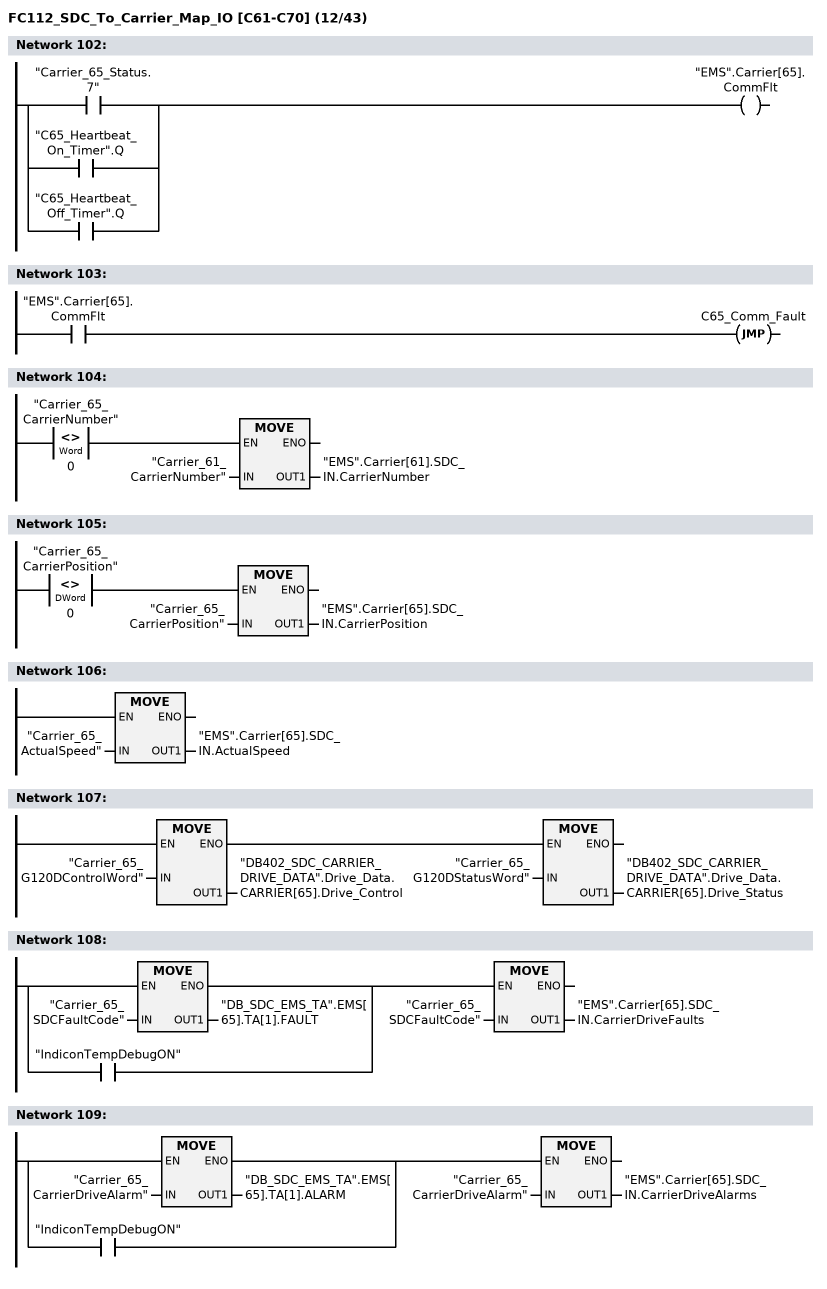
   RUNG wire#powerrail
      Contact( "Carrier_65_Status.7" )
      wire#w1
      Coil( "EMS".Carrier[65].CommFlt )
   END_RUNG
   RUNG wire#powerrail
      Contact( "C65_Heartbeat_On_Timer".Q )
   END_RUNG wire#w1
   RUNG wire#powerrail
      Contact( "C65_Heartbeat_Off_Timer".Q )
   END_RUNG wire#w1
   // the same network as SCL:
   "EMS".Carrier[65].CommFlt := "Carrier_65_Status.7" OR "C65_Heartbeat_On_Timer".Q OR "C65_Heartbeat_Off_Timer".Q;
END_REGION

REGION Network 103
   RUNG wire#powerrail
      Contact( "EMS".Carrier[65].CommFlt )
      JumpCoil( C65_Comm_Fault )
   END_RUNG
   // the same network as SCL:
   IF "EMS".Carrier[65].CommFlt THEN GOTO C65_Comm_Fault; END_IF;
END_REGION

REGION Network 104
   RUNG wire#powerrail
      { S7_Templates := "SrcType := Word" } NE_Contact(in1 := "Carrier_65_CarrierNumber", in2 := 0)
      Move(in := "Carrier_61_CarrierNumber", out1 => "EMS".Carrier[61].SDC_IN.CarrierNumber)
   END_RUNG
   // the same network as SCL:
   IF "Carrier_65_CarrierNumber" <> 0 THEN
       "EMS".Carrier[61].SDC_IN.CarrierNumber := "Carrier_61_CarrierNumber";
   END_IF;
END_REGION

REGION Network 105
   RUNG wire#powerrail
      { S7_Templates := "SrcType := DWord" } NE_Contact(in1 := "Carrier_65_CarrierPosition", in2 := 0)
      Move(in := "Carrier_65_CarrierPosition", out1 => "EMS".Carrier[65].SDC_IN.CarrierPosition)
   END_RUNG
   // the same network as SCL:
   IF "Carrier_65_CarrierPosition" <> 0 THEN
       "EMS".Carrier[65].SDC_IN.CarrierPosition := "Carrier_65_CarrierPosition";
   END_IF;
END_REGION

REGION Network 106
   RUNG wire#powerrail
      Move(in := "Carrier_65_ActualSpeed", out1 => "EMS".Carrier[65].SDC_IN.ActualSpeed)
   END_RUNG
   // the same network as SCL:
   "EMS".Carrier[65].SDC_IN.ActualSpeed := "Carrier_65_ActualSpeed";
END_REGION

REGION Network 107
   RUNG wire#powerrail
      Move(in := "Carrier_65_G120DControlWord", out1 => "DB402_SDC_CARRIER_DRIVE_DATA".Drive_Data.CARRIER[65].Drive_Control)
      Move(in := "Carrier_65_G120DStatusWord", out1 => "DB402_SDC_CARRIER_DRIVE_DATA".Drive_Data.CARRIER[65].Drive_Status)
   END_RUNG
   // the same network as SCL:
   "DB402_SDC_CARRIER_DRIVE_DATA".Drive_Data.CARRIER[65].Drive_Control := "Carrier_65_G120DControlWord";
   "DB402_SDC_CARRIER_DRIVE_DATA".Drive_Data.CARRIER[65].Drive_Status := "Carrier_65_G120DStatusWord";
END_REGION

REGION Network 108
   RUNG wire#powerrail
      Move(in := "Carrier_65_SDCFaultCode", out1 => "DB_SDC_EMS_TA".EMS[65].TA[1].FAULT)
      wire#w1
      Move(in := "Carrier_65_SDCFaultCode", out1 => "EMS".Carrier[65].SDC_IN.CarrierDriveFaults)
   END_RUNG
   RUNG wire#powerrail
      Contact( "IndiconTempDebugON" )
   END_RUNG wire#w1
   // the same network as SCL:
   "DB_SDC_EMS_TA".EMS[65].TA[1].FAULT := "Carrier_65_SDCFaultCode";
   IF TRUE OR "IndiconTempDebugON" THEN
       "EMS".Carrier[65].SDC_IN.CarrierDriveFaults := "Carrier_65_SDCFaultCode";
   END_IF;
END_REGION

REGION Network 109
   RUNG wire#powerrail
      Move(in := "Carrier_65_CarrierDriveAlarm", out1 => "DB_SDC_EMS_TA".EMS[65].TA[1].ALARM)
      wire#w1
      Move(in := "Carrier_65_CarrierDriveAlarm", out1 => "EMS".Carrier[65].SDC_IN.CarrierDriveAlarms)
   END_RUNG
   RUNG wire#powerrail
      Contact( "IndiconTempDebugON" )
   END_RUNG wire#w1
   // the same network as SCL:
   "DB_SDC_EMS_TA".EMS[65].TA[1].ALARM := "Carrier_65_CarrierDriveAlarm";
   IF TRUE OR "IndiconTempDebugON" THEN
       "EMS".Carrier[65].SDC_IN.CarrierDriveAlarms := "Carrier_65_CarrierDriveAlarm";
   END_IF;
END_REGION

REGION Network 110
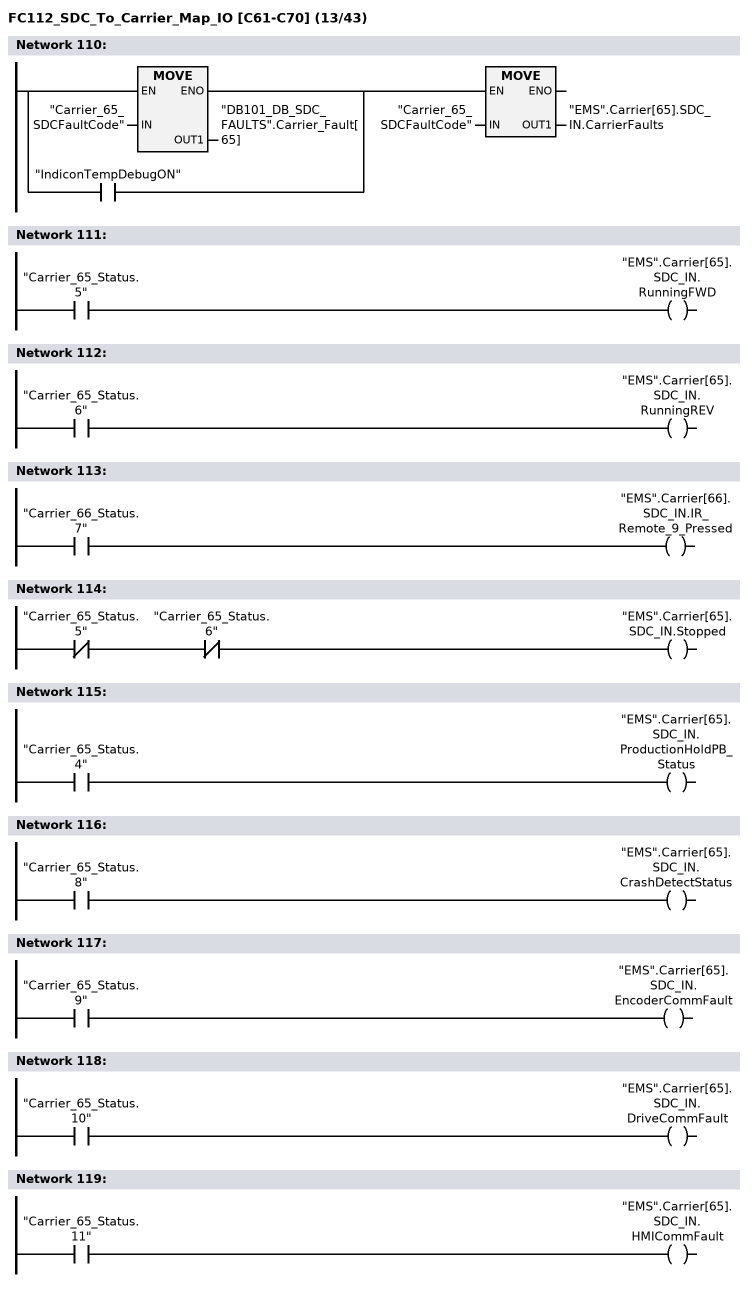
   RUNG wire#powerrail
      Move(in := "Carrier_65_SDCFaultCode", out1 => "DB101_DB_SDC_FAULTS".Carrier_Fault[65])
      wire#w1
      Move(in := "Carrier_65_SDCFaultCode", out1 => "EMS".Carrier[65].SDC_IN.CarrierFaults)
   END_RUNG
   RUNG wire#powerrail
      Contact( "IndiconTempDebugON" )
   END_RUNG wire#w1
   // the same network as SCL:
   "DB101_DB_SDC_FAULTS".Carrier_Fault[65] := "Carrier_65_SDCFaultCode";
   IF TRUE OR "IndiconTempDebugON" THEN
       "EMS".Carrier[65].SDC_IN.CarrierFaults := "Carrier_65_SDCFaultCode";
   END_IF;
END_REGION

REGION Network 111
   RUNG wire#powerrail
      Contact( "Carrier_65_Status.5" )
      Coil( "EMS".Carrier[65].SDC_IN.RunningFWD )
   END_RUNG
   // the same network as SCL:
   "EMS".Carrier[65].SDC_IN.RunningFWD := "Carrier_65_Status.5";
END_REGION

REGION Network 112
   RUNG wire#powerrail
      Contact( "Carrier_65_Status.6" )
      Coil( "EMS".Carrier[65].SDC_IN.RunningREV )
   END_RUNG
   // the same network as SCL:
   "EMS".Carrier[65].SDC_IN.RunningREV := "Carrier_65_Status.6";
END_REGION

REGION Network 113
   RUNG wire#powerrail
      Contact( "Carrier_66_Status.7" )
      Coil( "EMS".Carrier[66].SDC_IN.IR_Remote_9_Pressed )
   END_RUNG
   // the same network as SCL:
   "EMS".Carrier[66].SDC_IN.IR_Remote_9_Pressed := "Carrier_66_Status.7";
END_REGION

REGION Network 114
   RUNG wire#powerrail
      I_Contact( "Carrier_65_Status.5" )
      I_Contact( "Carrier_65_Status.6" )
      Coil( "EMS".Carrier[65].SDC_IN.Stopped )
   END_RUNG
   // the same network as SCL:
   "EMS".Carrier[65].SDC_IN.Stopped := NOT "Carrier_65_Status.5" AND NOT "Carrier_65_Status.6";
END_REGION

REGION Network 115
   RUNG wire#powerrail
      Contact( "Carrier_65_Status.4" )
      Coil( "EMS".Carrier[65].SDC_IN.ProductionHoldPB_Status )
   END_RUNG
   // the same network as SCL:
   "EMS".Carrier[65].SDC_IN.ProductionHoldPB_Status := "Carrier_65_Status.4";
END_REGION

REGION Network 116
   RUNG wire#powerrail
      Contact( "Carrier_65_Status.8" )
      Coil( "EMS".Carrier[65].SDC_IN.CrashDetectStatus )
   END_RUNG
   // the same network as SCL:
   "EMS".Carrier[65].SDC_IN.CrashDetectStatus := "Carrier_65_Status.8";
END_REGION

REGION Network 117
   RUNG wire#powerrail
      Contact( "Carrier_65_Status.9" )
      Coil( "EMS".Carrier[65].SDC_IN.EncoderCommFault )
   END_RUNG
   // the same network as SCL:
   "EMS".Carrier[65].SDC_IN.EncoderCommFault := "Carrier_65_Status.9";
END_REGION

REGION Network 118
   RUNG wire#powerrail
      Contact( "Carrier_65_Status.10" )
      Coil( "EMS".Carrier[65].SDC_IN.DriveCommFault )
   END_RUNG
   // the same network as SCL:
   "EMS".Carrier[65].SDC_IN.DriveCommFault := "Carrier_65_Status.10";
END_REGION

REGION Network 119
   RUNG wire#powerrail
      Contact( "Carrier_65_Status.11" )
      Coil( "EMS".Carrier[65].SDC_IN.HMICommFault )
   END_RUNG
   // the same network as SCL:
   "EMS".Carrier[65].SDC_IN.HMICommFault := "Carrier_65_Status.11";
END_REGION

REGION Network 120
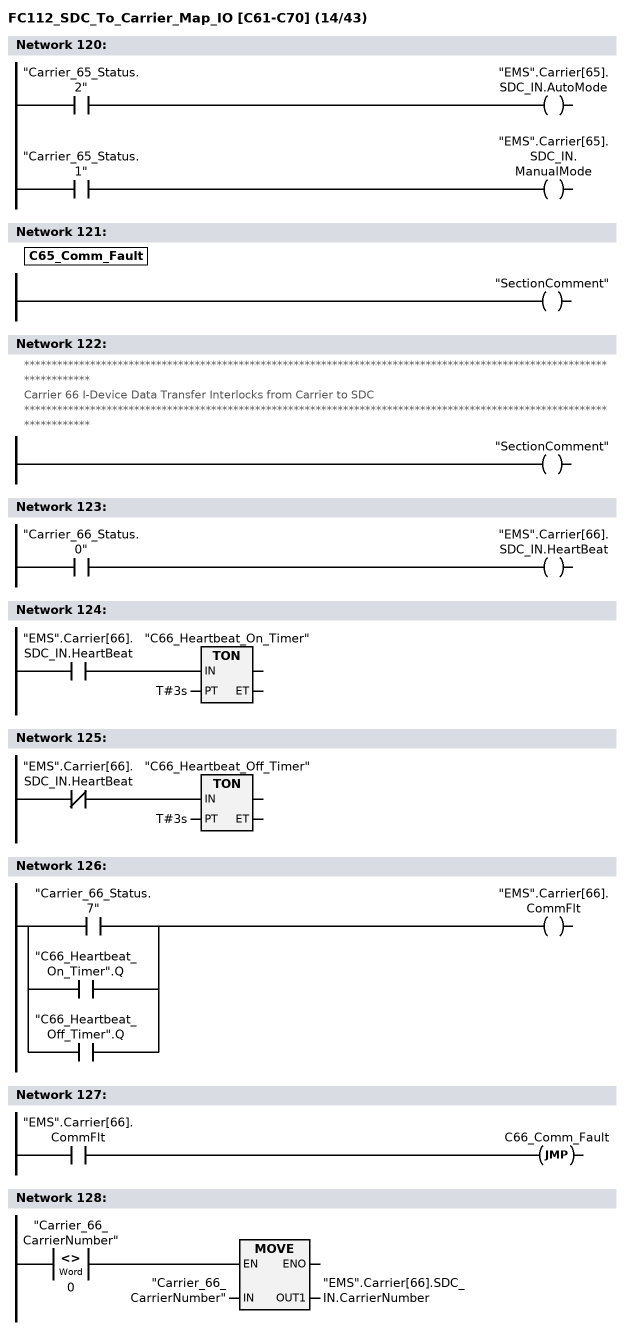
   RUNG wire#powerrail
      Contact( "Carrier_65_Status.2" )
      Coil( "EMS".Carrier[65].SDC_IN.AutoMode )
   END_RUNG
   RUNG wire#powerrail
      Contact( "Carrier_65_Status.1" )
      Coil( "EMS".Carrier[65].SDC_IN.ManualMode )
   END_RUNG
   // the same network as SCL:
   "EMS".Carrier[65].SDC_IN.AutoMode := "Carrier_65_Status.2";
   "EMS".Carrier[65].SDC_IN.ManualMode := "Carrier_65_Status.1";
END_REGION

REGION Network 121
   Label( C65_Comm_Fault )
   RUNG wire#powerrail
      Coil( "SectionComment" )
   END_RUNG
   // the same network as SCL:
   C65_Comm_Fault:
   "SectionComment" := TRUE;
END_REGION

REGION Network 122
   // **********************************************************************************************************************
   // 
   // Carrier 66 I-Device Data Transfer Interlocks from Carrier to SDC
   // 
   // **********************************************************************************************************************
   RUNG wire#powerrail
      Coil( "SectionComment" )
   END_RUNG
   // the same network as SCL:
   "SectionComment" := TRUE;
END_REGION

REGION Network 123
   RUNG wire#powerrail
      Contact( "Carrier_66_Status.0" )
      Coil( "EMS".Carrier[66].SDC_IN.HeartBeat )
   END_RUNG
   // the same network as SCL:
   "EMS".Carrier[66].SDC_IN.HeartBeat := "Carrier_66_Status.0";
END_REGION

REGION Network 124
   "C66_Heartbeat_On_Timer".TON(IN := "EMS".Carrier[66].SDC_IN.HeartBeat, PT := T#3s);
END_REGION

REGION Network 125
   "C66_Heartbeat_Off_Timer".TON(IN := NOT "EMS".Carrier[66].SDC_IN.HeartBeat, PT := T#3s);
END_REGION

REGION Network 126
   RUNG wire#powerrail
      Contact( "Carrier_66_Status.7" )
      wire#w1
      Coil( "EMS".Carrier[66].CommFlt )
   END_RUNG
   RUNG wire#powerrail
      Contact( "C66_Heartbeat_On_Timer".Q )
   END_RUNG wire#w1
   RUNG wire#powerrail
      Contact( "C66_Heartbeat_Off_Timer".Q )
   END_RUNG wire#w1
   // the same network as SCL:
   "EMS".Carrier[66].CommFlt := "Carrier_66_Status.7" OR "C66_Heartbeat_On_Timer".Q OR "C66_Heartbeat_Off_Timer".Q;
END_REGION

REGION Network 127
   RUNG wire#powerrail
      Contact( "EMS".Carrier[66].CommFlt )
      JumpCoil( C66_Comm_Fault )
   END_RUNG
   // the same network as SCL:
   IF "EMS".Carrier[66].CommFlt THEN GOTO C66_Comm_Fault; END_IF;
END_REGION

REGION Network 128
   RUNG wire#powerrail
      { S7_Templates := "SrcType := Word" } NE_Contact(in1 := "Carrier_66_CarrierNumber", in2 := 0)
      Move(in := "Carrier_66_CarrierNumber", out1 => "EMS".Carrier[66].SDC_IN.CarrierNumber)
   END_RUNG
   // the same network as SCL:
   IF "Carrier_66_CarrierNumber" <> 0 THEN
       "EMS".Carrier[66].SDC_IN.CarrierNumber := "Carrier_66_CarrierNumber";
   END_IF;
END_REGION

REGION Network 129
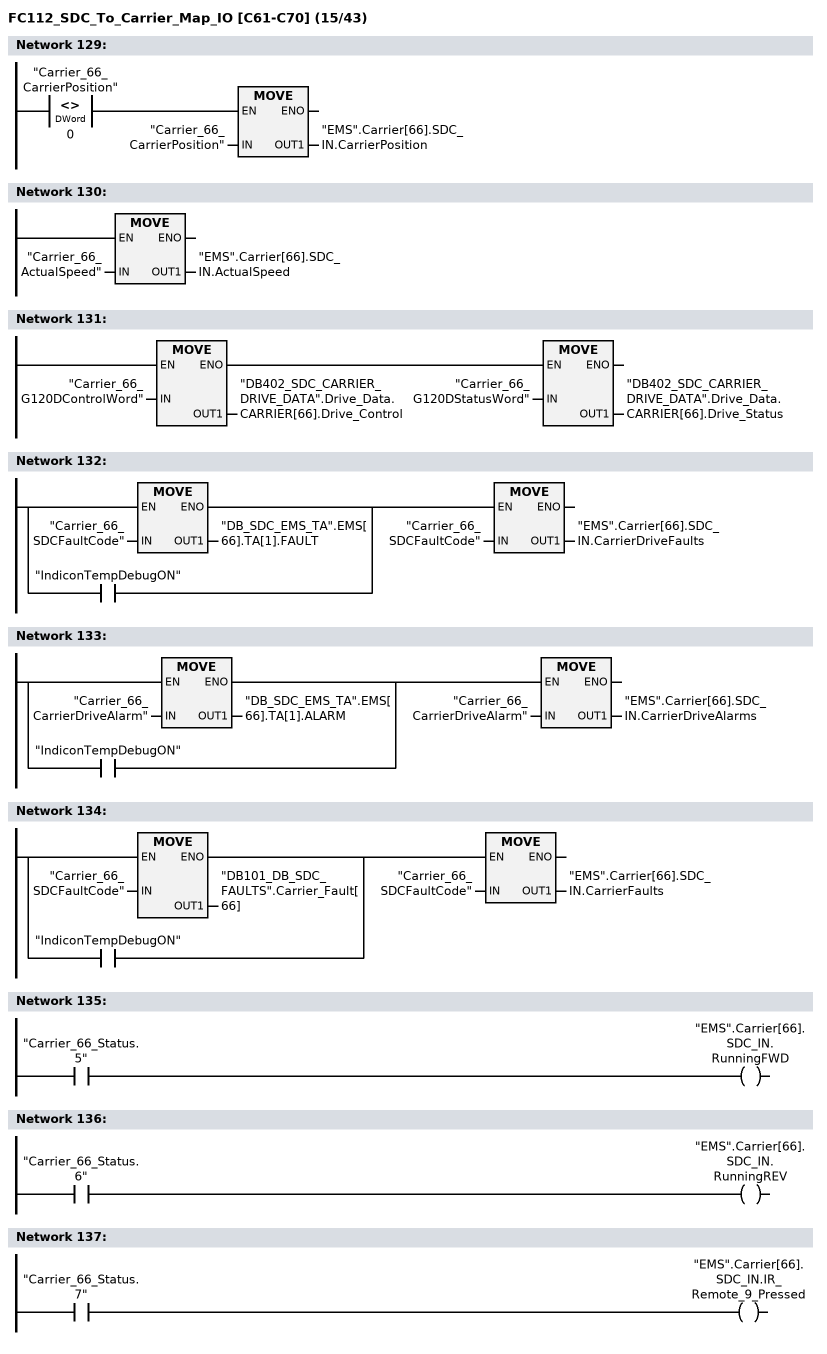
   RUNG wire#powerrail
      { S7_Templates := "SrcType := DWord" } NE_Contact(in1 := "Carrier_66_CarrierPosition", in2 := 0)
      Move(in := "Carrier_66_CarrierPosition", out1 => "EMS".Carrier[66].SDC_IN.CarrierPosition)
   END_RUNG
   // the same network as SCL:
   IF "Carrier_66_CarrierPosition" <> 0 THEN
       "EMS".Carrier[66].SDC_IN.CarrierPosition := "Carrier_66_CarrierPosition";
   END_IF;
END_REGION

REGION Network 130
   RUNG wire#powerrail
      Move(in := "Carrier_66_ActualSpeed", out1 => "EMS".Carrier[66].SDC_IN.ActualSpeed)
   END_RUNG
   // the same network as SCL:
   "EMS".Carrier[66].SDC_IN.ActualSpeed := "Carrier_66_ActualSpeed";
END_REGION

REGION Network 131
   RUNG wire#powerrail
      Move(in := "Carrier_66_G120DControlWord", out1 => "DB402_SDC_CARRIER_DRIVE_DATA".Drive_Data.CARRIER[66].Drive_Control)
      Move(in := "Carrier_66_G120DStatusWord", out1 => "DB402_SDC_CARRIER_DRIVE_DATA".Drive_Data.CARRIER[66].Drive_Status)
   END_RUNG
   // the same network as SCL:
   "DB402_SDC_CARRIER_DRIVE_DATA".Drive_Data.CARRIER[66].Drive_Control := "Carrier_66_G120DControlWord";
   "DB402_SDC_CARRIER_DRIVE_DATA".Drive_Data.CARRIER[66].Drive_Status := "Carrier_66_G120DStatusWord";
END_REGION

REGION Network 132
   RUNG wire#powerrail
      Move(in := "Carrier_66_SDCFaultCode", out1 => "DB_SDC_EMS_TA".EMS[66].TA[1].FAULT)
      wire#w1
      Move(in := "Carrier_66_SDCFaultCode", out1 => "EMS".Carrier[66].SDC_IN.CarrierDriveFaults)
   END_RUNG
   RUNG wire#powerrail
      Contact( "IndiconTempDebugON" )
   END_RUNG wire#w1
   // the same network as SCL:
   "DB_SDC_EMS_TA".EMS[66].TA[1].FAULT := "Carrier_66_SDCFaultCode";
   IF TRUE OR "IndiconTempDebugON" THEN
       "EMS".Carrier[66].SDC_IN.CarrierDriveFaults := "Carrier_66_SDCFaultCode";
   END_IF;
END_REGION

REGION Network 133
   RUNG wire#powerrail
      Move(in := "Carrier_66_CarrierDriveAlarm", out1 => "DB_SDC_EMS_TA".EMS[66].TA[1].ALARM)
      wire#w1
      Move(in := "Carrier_66_CarrierDriveAlarm", out1 => "EMS".Carrier[66].SDC_IN.CarrierDriveAlarms)
   END_RUNG
   RUNG wire#powerrail
      Contact( "IndiconTempDebugON" )
   END_RUNG wire#w1
   // the same network as SCL:
   "DB_SDC_EMS_TA".EMS[66].TA[1].ALARM := "Carrier_66_CarrierDriveAlarm";
   IF TRUE OR "IndiconTempDebugON" THEN
       "EMS".Carrier[66].SDC_IN.CarrierDriveAlarms := "Carrier_66_CarrierDriveAlarm";
   END_IF;
END_REGION

REGION Network 134
   RUNG wire#powerrail
      Move(in := "Carrier_66_SDCFaultCode", out1 => "DB101_DB_SDC_FAULTS".Carrier_Fault[66])
      wire#w1
      Move(in := "Carrier_66_SDCFaultCode", out1 => "EMS".Carrier[66].SDC_IN.CarrierFaults)
   END_RUNG
   RUNG wire#powerrail
      Contact( "IndiconTempDebugON" )
   END_RUNG wire#w1
   // the same network as SCL:
   "DB101_DB_SDC_FAULTS".Carrier_Fault[66] := "Carrier_66_SDCFaultCode";
   IF TRUE OR "IndiconTempDebugON" THEN
       "EMS".Carrier[66].SDC_IN.CarrierFaults := "Carrier_66_SDCFaultCode";
   END_IF;
END_REGION

REGION Network 135
   RUNG wire#powerrail
      Contact( "Carrier_66_Status.5" )
      Coil( "EMS".Carrier[66].SDC_IN.RunningFWD )
   END_RUNG
   // the same network as SCL:
   "EMS".Carrier[66].SDC_IN.RunningFWD := "Carrier_66_Status.5";
END_REGION

REGION Network 136
   RUNG wire#powerrail
      Contact( "Carrier_66_Status.6" )
      Coil( "EMS".Carrier[66].SDC_IN.RunningREV )
   END_RUNG
   // the same network as SCL:
   "EMS".Carrier[66].SDC_IN.RunningREV := "Carrier_66_Status.6";
END_REGION

REGION Network 137
   RUNG wire#powerrail
      Contact( "Carrier_66_Status.7" )
      Coil( "EMS".Carrier[66].SDC_IN.IR_Remote_9_Pressed )
   END_RUNG
   // the same network as SCL:
   "EMS".Carrier[66].SDC_IN.IR_Remote_9_Pressed := "Carrier_66_Status.7";
END_REGION

REGION Network 138
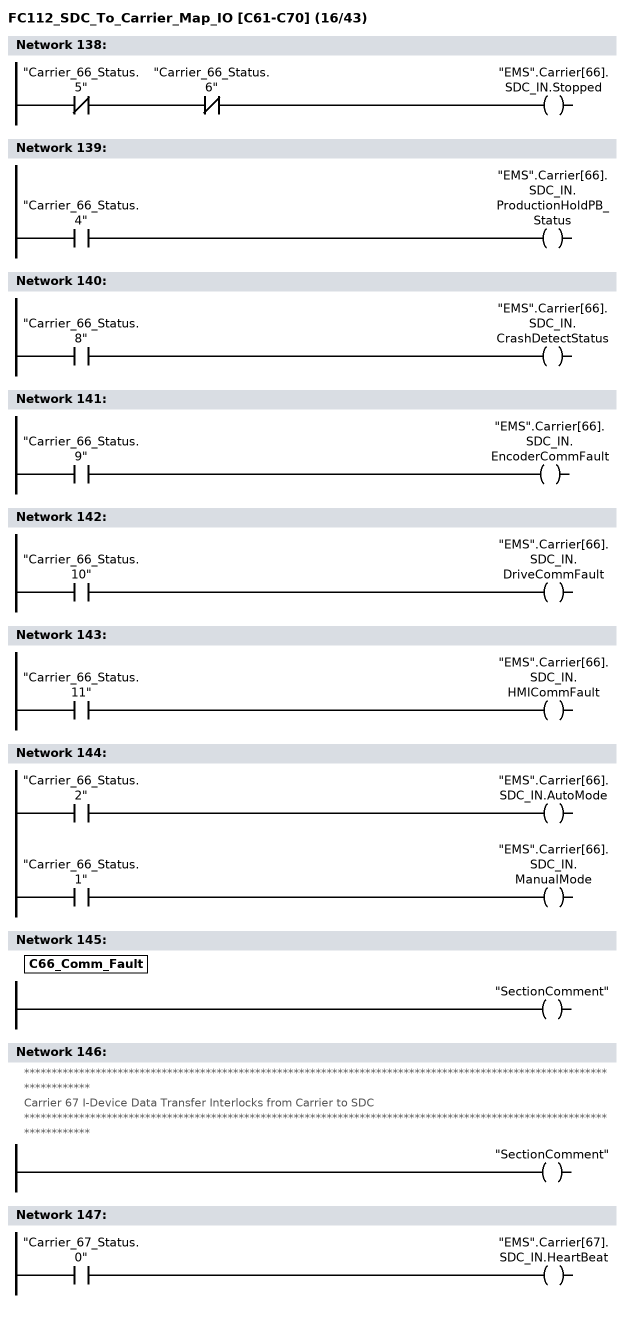
   RUNG wire#powerrail
      I_Contact( "Carrier_66_Status.5" )
      I_Contact( "Carrier_66_Status.6" )
      Coil( "EMS".Carrier[66].SDC_IN.Stopped )
   END_RUNG
   // the same network as SCL:
   "EMS".Carrier[66].SDC_IN.Stopped := NOT "Carrier_66_Status.5" AND NOT "Carrier_66_Status.6";
END_REGION

REGION Network 139
   RUNG wire#powerrail
      Contact( "Carrier_66_Status.4" )
      Coil( "EMS".Carrier[66].SDC_IN.ProductionHoldPB_Status )
   END_RUNG
   // the same network as SCL:
   "EMS".Carrier[66].SDC_IN.ProductionHoldPB_Status := "Carrier_66_Status.4";
END_REGION

REGION Network 140
   RUNG wire#powerrail
      Contact( "Carrier_66_Status.8" )
      Coil( "EMS".Carrier[66].SDC_IN.CrashDetectStatus )
   END_RUNG
   // the same network as SCL:
   "EMS".Carrier[66].SDC_IN.CrashDetectStatus := "Carrier_66_Status.8";
END_REGION

REGION Network 141
   RUNG wire#powerrail
      Contact( "Carrier_66_Status.9" )
      Coil( "EMS".Carrier[66].SDC_IN.EncoderCommFault )
   END_RUNG
   // the same network as SCL:
   "EMS".Carrier[66].SDC_IN.EncoderCommFault := "Carrier_66_Status.9";
END_REGION

REGION Network 142
   RUNG wire#powerrail
      Contact( "Carrier_66_Status.10" )
      Coil( "EMS".Carrier[66].SDC_IN.DriveCommFault )
   END_RUNG
   // the same network as SCL:
   "EMS".Carrier[66].SDC_IN.DriveCommFault := "Carrier_66_Status.10";
END_REGION

REGION Network 143
   RUNG wire#powerrail
      Contact( "Carrier_66_Status.11" )
      Coil( "EMS".Carrier[66].SDC_IN.HMICommFault )
   END_RUNG
   // the same network as SCL:
   "EMS".Carrier[66].SDC_IN.HMICommFault := "Carrier_66_Status.11";
END_REGION

REGION Network 144
   RUNG wire#powerrail
      Contact( "Carrier_66_Status.2" )
      Coil( "EMS".Carrier[66].SDC_IN.AutoMode )
   END_RUNG
   RUNG wire#powerrail
      Contact( "Carrier_66_Status.1" )
      Coil( "EMS".Carrier[66].SDC_IN.ManualMode )
   END_RUNG
   // the same network as SCL:
   "EMS".Carrier[66].SDC_IN.AutoMode := "Carrier_66_Status.2";
   "EMS".Carrier[66].SDC_IN.ManualMode := "Carrier_66_Status.1";
END_REGION

REGION Network 145
   Label( C66_Comm_Fault )
   RUNG wire#powerrail
      Coil( "SectionComment" )
   END_RUNG
   // the same network as SCL:
   C66_Comm_Fault:
   "SectionComment" := TRUE;
END_REGION

REGION Network 146
   // **********************************************************************************************************************
   // 
   // Carrier 67 I-Device Data Transfer Interlocks from Carrier to SDC
   // 
   // **********************************************************************************************************************
   RUNG wire#powerrail
      Coil( "SectionComment" )
   END_RUNG
   // the same network as SCL:
   "SectionComment" := TRUE;
END_REGION

REGION Network 147
   RUNG wire#powerrail
      Contact( "Carrier_67_Status.0" )
      Coil( "EMS".Carrier[67].SDC_IN.HeartBeat )
   END_RUNG
   // the same network as SCL:
   "EMS".Carrier[67].SDC_IN.HeartBeat := "Carrier_67_Status.0";
END_REGION

REGION Network 148
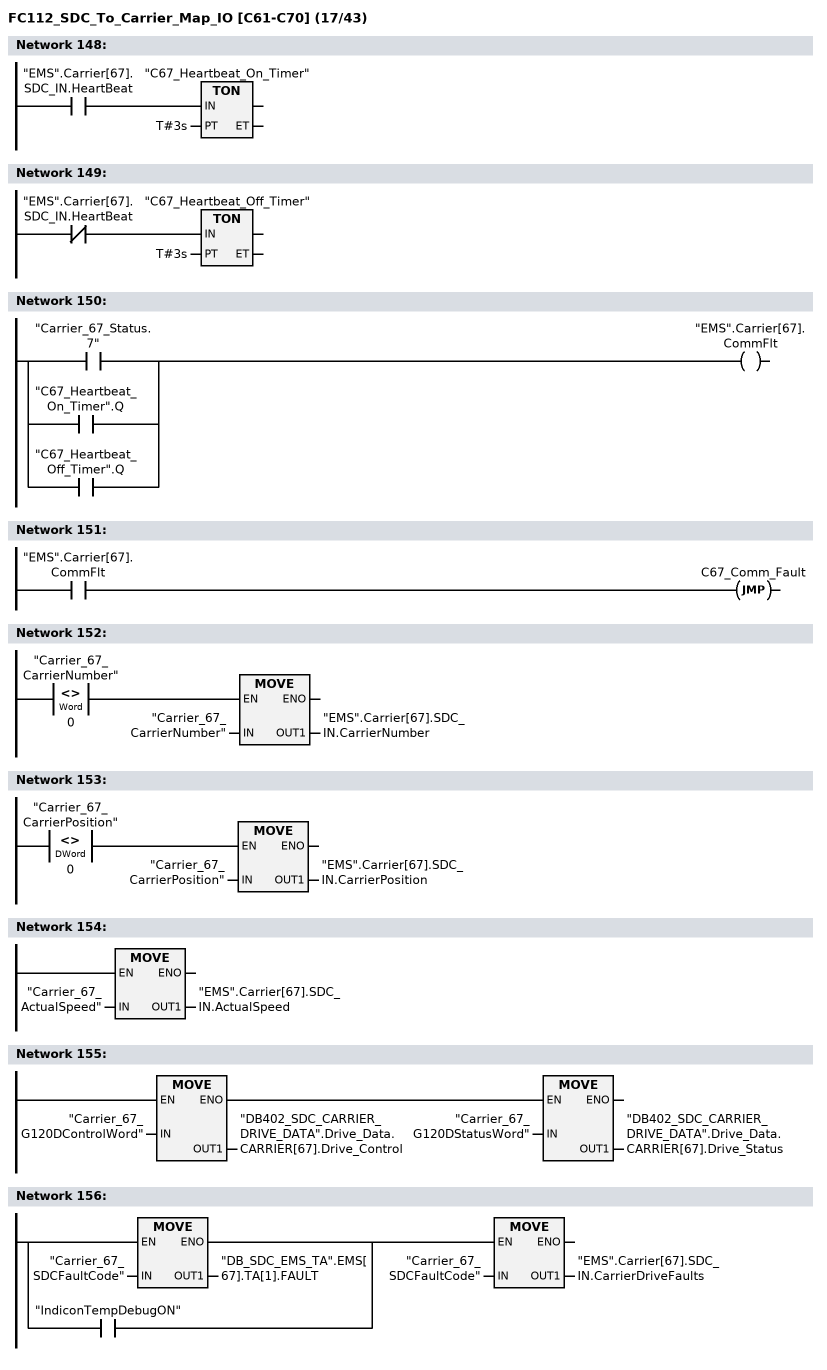
   "C67_Heartbeat_On_Timer".TON(IN := "EMS".Carrier[67].SDC_IN.HeartBeat, PT := T#3s);
END_REGION

REGION Network 149
   "C67_Heartbeat_Off_Timer".TON(IN := NOT "EMS".Carrier[67].SDC_IN.HeartBeat, PT := T#3s);
END_REGION

REGION Network 150
   RUNG wire#powerrail
      Contact( "Carrier_67_Status.7" )
      wire#w1
      Coil( "EMS".Carrier[67].CommFlt )
   END_RUNG
   RUNG wire#powerrail
      Contact( "C67_Heartbeat_On_Timer".Q )
   END_RUNG wire#w1
   RUNG wire#powerrail
      Contact( "C67_Heartbeat_Off_Timer".Q )
   END_RUNG wire#w1
   // the same network as SCL:
   "EMS".Carrier[67].CommFlt := "Carrier_67_Status.7" OR "C67_Heartbeat_On_Timer".Q OR "C67_Heartbeat_Off_Timer".Q;
END_REGION

REGION Network 151
   RUNG wire#powerrail
      Contact( "EMS".Carrier[67].CommFlt )
      JumpCoil( C67_Comm_Fault )
   END_RUNG
   // the same network as SCL:
   IF "EMS".Carrier[67].CommFlt THEN GOTO C67_Comm_Fault; END_IF;
END_REGION

REGION Network 152
   RUNG wire#powerrail
      { S7_Templates := "SrcType := Word" } NE_Contact(in1 := "Carrier_67_CarrierNumber", in2 := 0)
      Move(in := "Carrier_67_CarrierNumber", out1 => "EMS".Carrier[67].SDC_IN.CarrierNumber)
   END_RUNG
   // the same network as SCL:
   IF "Carrier_67_CarrierNumber" <> 0 THEN
       "EMS".Carrier[67].SDC_IN.CarrierNumber := "Carrier_67_CarrierNumber";
   END_IF;
END_REGION

REGION Network 153
   RUNG wire#powerrail
      { S7_Templates := "SrcType := DWord" } NE_Contact(in1 := "Carrier_67_CarrierPosition", in2 := 0)
      Move(in := "Carrier_67_CarrierPosition", out1 => "EMS".Carrier[67].SDC_IN.CarrierPosition)
   END_RUNG
   // the same network as SCL:
   IF "Carrier_67_CarrierPosition" <> 0 THEN
       "EMS".Carrier[67].SDC_IN.CarrierPosition := "Carrier_67_CarrierPosition";
   END_IF;
END_REGION

REGION Network 154
   RUNG wire#powerrail
      Move(in := "Carrier_67_ActualSpeed", out1 => "EMS".Carrier[67].SDC_IN.ActualSpeed)
   END_RUNG
   // the same network as SCL:
   "EMS".Carrier[67].SDC_IN.ActualSpeed := "Carrier_67_ActualSpeed";
END_REGION

REGION Network 155
   RUNG wire#powerrail
      Move(in := "Carrier_67_G120DControlWord", out1 => "DB402_SDC_CARRIER_DRIVE_DATA".Drive_Data.CARRIER[67].Drive_Control)
      Move(in := "Carrier_67_G120DStatusWord", out1 => "DB402_SDC_CARRIER_DRIVE_DATA".Drive_Data.CARRIER[67].Drive_Status)
   END_RUNG
   // the same network as SCL:
   "DB402_SDC_CARRIER_DRIVE_DATA".Drive_Data.CARRIER[67].Drive_Control := "Carrier_67_G120DControlWord";
   "DB402_SDC_CARRIER_DRIVE_DATA".Drive_Data.CARRIER[67].Drive_Status := "Carrier_67_G120DStatusWord";
END_REGION

REGION Network 156
   RUNG wire#powerrail
      Move(in := "Carrier_67_SDCFaultCode", out1 => "DB_SDC_EMS_TA".EMS[67].TA[1].FAULT)
      wire#w1
      Move(in := "Carrier_67_SDCFaultCode", out1 => "EMS".Carrier[67].SDC_IN.CarrierDriveFaults)
   END_RUNG
   RUNG wire#powerrail
      Contact( "IndiconTempDebugON" )
   END_RUNG wire#w1
   // the same network as SCL:
   "DB_SDC_EMS_TA".EMS[67].TA[1].FAULT := "Carrier_67_SDCFaultCode";
   IF TRUE OR "IndiconTempDebugON" THEN
       "EMS".Carrier[67].SDC_IN.CarrierDriveFaults := "Carrier_67_SDCFaultCode";
   END_IF;
END_REGION

REGION Network 157
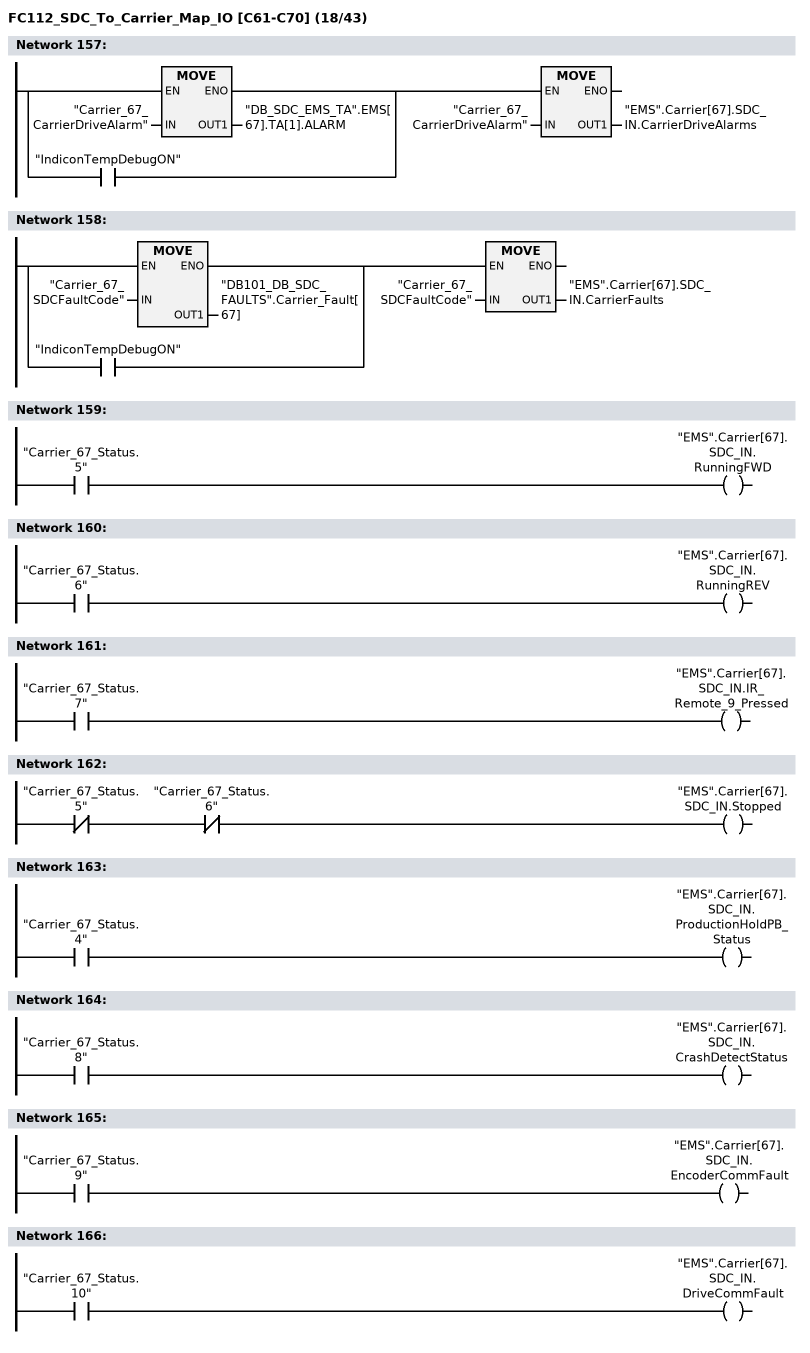
   RUNG wire#powerrail
      Move(in := "Carrier_67_CarrierDriveAlarm", out1 => "DB_SDC_EMS_TA".EMS[67].TA[1].ALARM)
      wire#w1
      Move(in := "Carrier_67_CarrierDriveAlarm", out1 => "EMS".Carrier[67].SDC_IN.CarrierDriveAlarms)
   END_RUNG
   RUNG wire#powerrail
      Contact( "IndiconTempDebugON" )
   END_RUNG wire#w1
   // the same network as SCL:
   "DB_SDC_EMS_TA".EMS[67].TA[1].ALARM := "Carrier_67_CarrierDriveAlarm";
   IF TRUE OR "IndiconTempDebugON" THEN
       "EMS".Carrier[67].SDC_IN.CarrierDriveAlarms := "Carrier_67_CarrierDriveAlarm";
   END_IF;
END_REGION

REGION Network 158
   RUNG wire#powerrail
      Move(in := "Carrier_67_SDCFaultCode", out1 => "DB101_DB_SDC_FAULTS".Carrier_Fault[67])
      wire#w1
      Move(in := "Carrier_67_SDCFaultCode", out1 => "EMS".Carrier[67].SDC_IN.CarrierFaults)
   END_RUNG
   RUNG wire#powerrail
      Contact( "IndiconTempDebugON" )
   END_RUNG wire#w1
   // the same network as SCL:
   "DB101_DB_SDC_FAULTS".Carrier_Fault[67] := "Carrier_67_SDCFaultCode";
   IF TRUE OR "IndiconTempDebugON" THEN
       "EMS".Carrier[67].SDC_IN.CarrierFaults := "Carrier_67_SDCFaultCode";
   END_IF;
END_REGION

REGION Network 159
   RUNG wire#powerrail
      Contact( "Carrier_67_Status.5" )
      Coil( "EMS".Carrier[67].SDC_IN.RunningFWD )
   END_RUNG
   // the same network as SCL:
   "EMS".Carrier[67].SDC_IN.RunningFWD := "Carrier_67_Status.5";
END_REGION

REGION Network 160
   RUNG wire#powerrail
      Contact( "Carrier_67_Status.6" )
      Coil( "EMS".Carrier[67].SDC_IN.RunningREV )
   END_RUNG
   // the same network as SCL:
   "EMS".Carrier[67].SDC_IN.RunningREV := "Carrier_67_Status.6";
END_REGION

REGION Network 161
   RUNG wire#powerrail
      Contact( "Carrier_67_Status.7" )
      Coil( "EMS".Carrier[67].SDC_IN.IR_Remote_9_Pressed )
   END_RUNG
   // the same network as SCL:
   "EMS".Carrier[67].SDC_IN.IR_Remote_9_Pressed := "Carrier_67_Status.7";
END_REGION

REGION Network 162
   RUNG wire#powerrail
      I_Contact( "Carrier_67_Status.5" )
      I_Contact( "Carrier_67_Status.6" )
      Coil( "EMS".Carrier[67].SDC_IN.Stopped )
   END_RUNG
   // the same network as SCL:
   "EMS".Carrier[67].SDC_IN.Stopped := NOT "Carrier_67_Status.5" AND NOT "Carrier_67_Status.6";
END_REGION

REGION Network 163
   RUNG wire#powerrail
      Contact( "Carrier_67_Status.4" )
      Coil( "EMS".Carrier[67].SDC_IN.ProductionHoldPB_Status )
   END_RUNG
   // the same network as SCL:
   "EMS".Carrier[67].SDC_IN.ProductionHoldPB_Status := "Carrier_67_Status.4";
END_REGION

REGION Network 164
   RUNG wire#powerrail
      Contact( "Carrier_67_Status.8" )
      Coil( "EMS".Carrier[67].SDC_IN.CrashDetectStatus )
   END_RUNG
   // the same network as SCL:
   "EMS".Carrier[67].SDC_IN.CrashDetectStatus := "Carrier_67_Status.8";
END_REGION

REGION Network 165
   RUNG wire#powerrail
      Contact( "Carrier_67_Status.9" )
      Coil( "EMS".Carrier[67].SDC_IN.EncoderCommFault )
   END_RUNG
   // the same network as SCL:
   "EMS".Carrier[67].SDC_IN.EncoderCommFault := "Carrier_67_Status.9";
END_REGION

REGION Network 166
   RUNG wire#powerrail
      Contact( "Carrier_67_Status.10" )
      Coil( "EMS".Carrier[67].SDC_IN.DriveCommFault )
   END_RUNG
   // the same network as SCL:
   "EMS".Carrier[67].SDC_IN.DriveCommFault := "Carrier_67_Status.10";
END_REGION

REGION Network 167
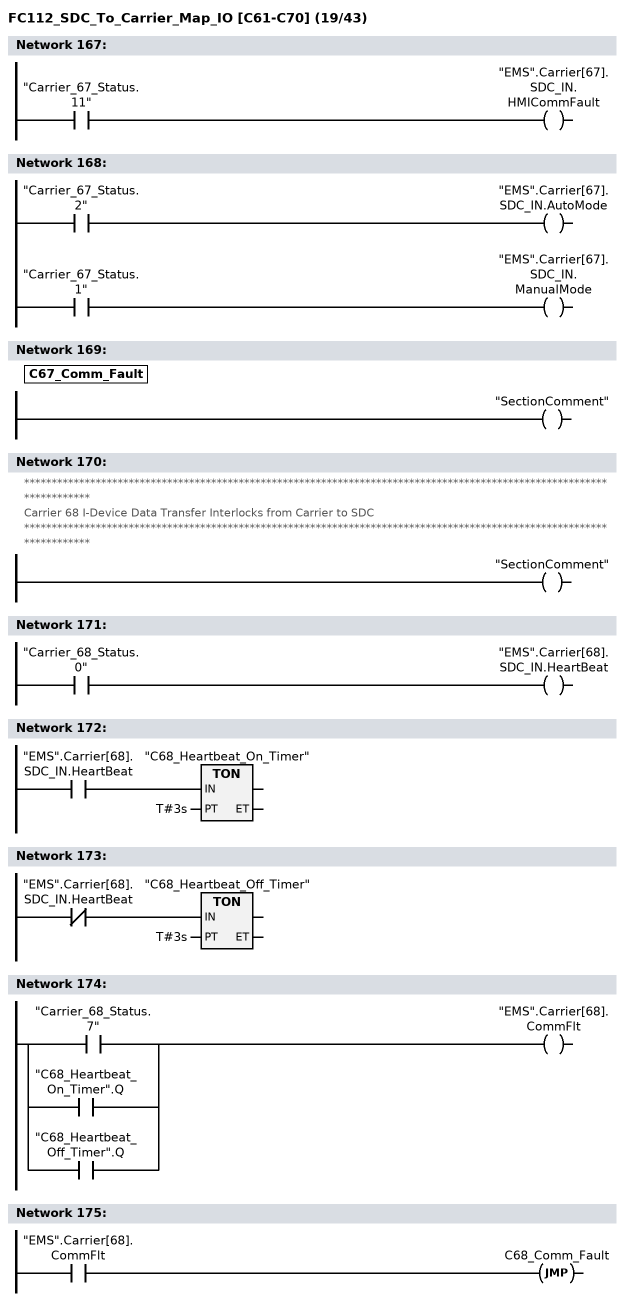
   RUNG wire#powerrail
      Contact( "Carrier_67_Status.11" )
      Coil( "EMS".Carrier[67].SDC_IN.HMICommFault )
   END_RUNG
   // the same network as SCL:
   "EMS".Carrier[67].SDC_IN.HMICommFault := "Carrier_67_Status.11";
END_REGION

REGION Network 168
   RUNG wire#powerrail
      Contact( "Carrier_67_Status.2" )
      Coil( "EMS".Carrier[67].SDC_IN.AutoMode )
   END_RUNG
   RUNG wire#powerrail
      Contact( "Carrier_67_Status.1" )
      Coil( "EMS".Carrier[67].SDC_IN.ManualMode )
   END_RUNG
   // the same network as SCL:
   "EMS".Carrier[67].SDC_IN.AutoMode := "Carrier_67_Status.2";
   "EMS".Carrier[67].SDC_IN.ManualMode := "Carrier_67_Status.1";
END_REGION

REGION Network 169
   Label( C67_Comm_Fault )
   RUNG wire#powerrail
      Coil( "SectionComment" )
   END_RUNG
   // the same network as SCL:
   C67_Comm_Fault:
   "SectionComment" := TRUE;
END_REGION

REGION Network 170
   // **********************************************************************************************************************
   // 
   // Carrier 68 I-Device Data Transfer Interlocks from Carrier to SDC
   // 
   // **********************************************************************************************************************
   RUNG wire#powerrail
      Coil( "SectionComment" )
   END_RUNG
   // the same network as SCL:
   "SectionComment" := TRUE;
END_REGION

REGION Network 171
   RUNG wire#powerrail
      Contact( "Carrier_68_Status.0" )
      Coil( "EMS".Carrier[68].SDC_IN.HeartBeat )
   END_RUNG
   // the same network as SCL:
   "EMS".Carrier[68].SDC_IN.HeartBeat := "Carrier_68_Status.0";
END_REGION

REGION Network 172
   "C68_Heartbeat_On_Timer".TON(IN := "EMS".Carrier[68].SDC_IN.HeartBeat, PT := T#3s);
END_REGION

REGION Network 173
   "C68_Heartbeat_Off_Timer".TON(IN := NOT "EMS".Carrier[68].SDC_IN.HeartBeat, PT := T#3s);
END_REGION

REGION Network 174
   RUNG wire#powerrail
      Contact( "Carrier_68_Status.7" )
      wire#w1
      Coil( "EMS".Carrier[68].CommFlt )
   END_RUNG
   RUNG wire#powerrail
      Contact( "C68_Heartbeat_On_Timer".Q )
   END_RUNG wire#w1
   RUNG wire#powerrail
      Contact( "C68_Heartbeat_Off_Timer".Q )
   END_RUNG wire#w1
   // the same network as SCL:
   "EMS".Carrier[68].CommFlt := "Carrier_68_Status.7" OR "C68_Heartbeat_On_Timer".Q OR "C68_Heartbeat_Off_Timer".Q;
END_REGION
